// TIA Portal project "e045002v087-088" (V13) (continued)
VERSION : 0.1
// stored: InstanceOfName FB_CTR_VAL
"FB_CTR_VAL"
BEGIN
END_DATA_BLOCK

DATA_BLOCK "STOP_PALLET"   // DB78
{ S7_Optimized_Access := 'FALSE' }
VERSION : 0.1
// stored: InstanceOfName FB_CTR_VAL
"FB_CTR_VAL"
BEGIN
END_DATA_BLOCK

DATA_BLOCK "FB_CTR_MOT_FRD_DB"   // DB104
{ S7_Optimized_Access := 'FALSE' }
VERSION : 0.1
// stored: InstanceOfName FB_CTR_MOT_FRD
"FB_CTR_MOT_FRD"
BEGIN
END_DATA_BLOCK

DATA_BLOCK "FB_CTR_MOT_FRD_DB_1"   // DB109
{ S7_Optimized_Access := 'FALSE' }
VERSION : 0.1
// stored: InstanceOfName FB_CTR_MOT_FRD
"FB_CTR_MOT_FRD"
BEGIN
END_DATA_BLOCK

DATA_BLOCK "FB_CTR_MOT_FRD_DB_2"   // DB145
{ S7_Optimized_Access := 'FALSE' }
VERSION : 0.1
// stored: InstanceOfName FB_CTR_MOT_FRD
"FB_CTR_MOT_FRD"
BEGIN
END_DATA_BLOCK

// folder: Movimiento DATOS

DATA_BLOCK "DB_RECETAS"   // DB4
{ S7_Optimized_Access := 'FALSE' }
VERSION : 0.1
   VAR
      Receta : Array [1..10] of "Recetas";
      Static_1 : Bool;
   END_VAR
BEGIN
END_DATA_BLOCK

DATA_BLOCK "Puntero"   // DB7
{ S7_Optimized_Access := 'FALSE' }
VERSION : 0.1
   VAR
      Max_Nro_Elementos : Word;
      Max_Nro_Filas : Word;
      Max_Nro_Capas : Word;
      Max_Nro_Recetas : Word;
      Offset_Filas_HMI : Word;
      Length_Filas_HMI : Word;
      Offset_Elementos_HMI : Word;
      Length_Elementos_HMI : Word;
      Offset_Recetas : Word;
      Length_Recetas : Word;
      Offset_Nombre_Receta : Word;
      Length_Nombre_Receta : Word;
      Offset_CantCapas_Receta : Word;
      Offset_CapasDist_Receta : Word;
      Offset_Capas_Receta : Word;
      Length_Capas_Receta : Word;
      Offset_Filas_CapaReceta : Word;
      Length_Filas_CapaReceta : Word;
      Offset_Vel_Dosificador : Word;
      Length_Vel_Dosificador : Word;
   END_VAR
BEGIN
END_DATA_BLOCK

DATA_BLOCK "DB_Receta_Actual"   // DB42
{ S7_Optimized_Access := 'FALSE' }
VERSION : 0.1
   VAR
      Número : Byte;
      Nombre : Array [1 .. 50] of Char;
      Nro_Capas_Pallet : Byte;
      Nro_Capas_Distintas : Byte;
      Capa : Array [1..10] of "Capas_Proceso";
      Static_1 : Bool;
   END_VAR
BEGIN
END_DATA_BLOCK

// folder: (top level)

FUNCTION "Valida_Velocidades" : Void   // FC2, LAD
{ S7_Optimized_Access := 'FALSE' }
VERSION : 0.1
BEGIN

REGION Network 1: Dosificador
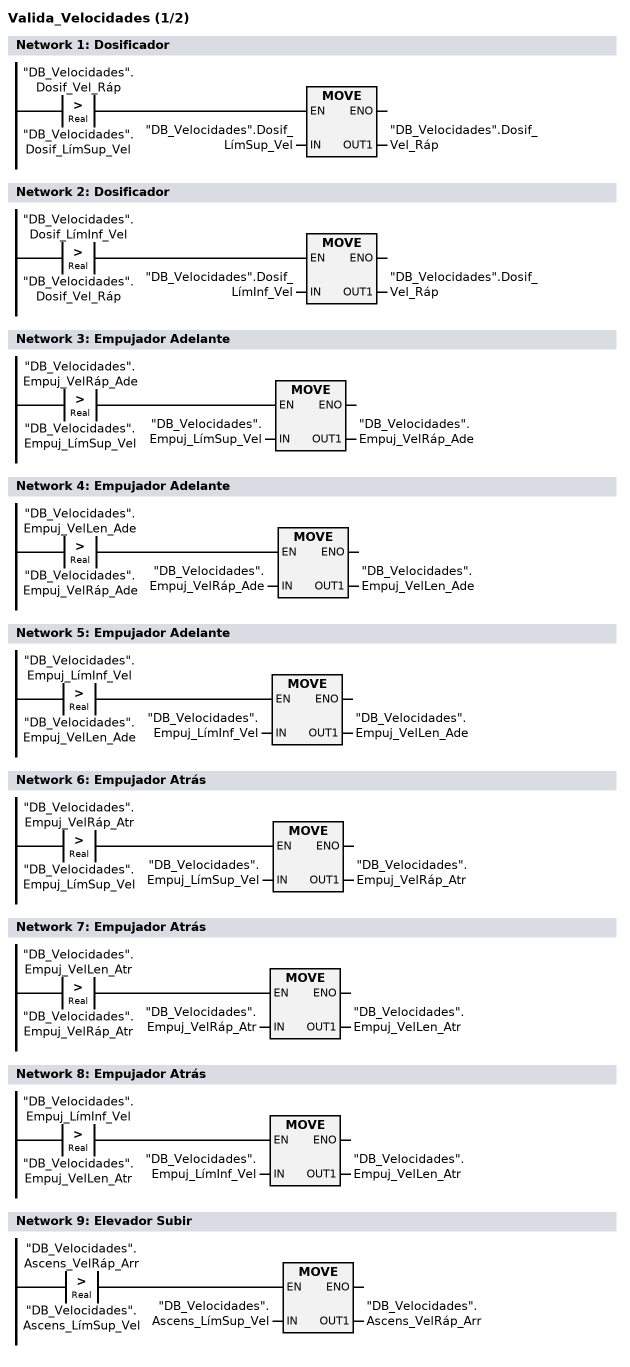
   RUNG wire#powerrail
      { S7_Templates := "SrcType := Real" } GT_Contact(in1 := "DB_Velocidades".Dosif_Vel_Ráp, in2 := "DB_Velocidades".Dosif_LímSup_Vel)
      { S7_GenerateENO := "TRUE" } Move(in := "DB_Velocidades".Dosif_LímSup_Vel, out1 => "DB_Velocidades".Dosif_Vel_Ráp)
   END_RUNG
   // the same network as SCL:
   IF "DB_Velocidades".Dosif_Vel_Ráp > "DB_Velocidades".Dosif_LímSup_Vel THEN
       "DB_Velocidades".Dosif_Vel_Ráp := "DB_Velocidades".Dosif_LímSup_Vel;
   END_IF;
END_REGION

REGION Network 2: Dosificador
   RUNG wire#powerrail
      { S7_Templates := "SrcType := Real" } GT_Contact(in1 := "DB_Velocidades".Dosif_LímInf_Vel, in2 := "DB_Velocidades".Dosif_Vel_Ráp)
      { S7_GenerateENO := "TRUE" } Move(in := "DB_Velocidades".Dosif_LímInf_Vel, out1 => "DB_Velocidades".Dosif_Vel_Ráp)
   END_RUNG
   // the same network as SCL:
   IF "DB_Velocidades".Dosif_LímInf_Vel > "DB_Velocidades".Dosif_Vel_Ráp THEN
       "DB_Velocidades".Dosif_Vel_Ráp := "DB_Velocidades".Dosif_LímInf_Vel;
   END_IF;
END_REGION

REGION Network 3: Empujador Adelante
   RUNG wire#powerrail
      { S7_Templates := "SrcType := Real" } GT_Contact(in1 := "DB_Velocidades".Empuj_VelRáp_Ade, in2 := "DB_Velocidades".Empuj_LímSup_Vel)
      { S7_GenerateENO := "TRUE" } Move(in := "DB_Velocidades".Empuj_LímSup_Vel, out1 => "DB_Velocidades".Empuj_VelRáp_Ade)
   END_RUNG
   // the same network as SCL:
   IF "DB_Velocidades".Empuj_VelRáp_Ade > "DB_Velocidades".Empuj_LímSup_Vel THEN
       "DB_Velocidades".Empuj_VelRáp_Ade := "DB_Velocidades".Empuj_LímSup_Vel;
   END_IF;
END_REGION

REGION Network 4: Empujador Adelante
   RUNG wire#powerrail
      { S7_Templates := "SrcType := Real" } GT_Contact(in1 := "DB_Velocidades".Empuj_VelLen_Ade, in2 := "DB_Velocidades".Empuj_VelRáp_Ade)
      { S7_GenerateENO := "TRUE" } Move(in := "DB_Velocidades".Empuj_VelRáp_Ade, out1 => "DB_Velocidades".Empuj_VelLen_Ade)
   END_RUNG
   // the same network as SCL:
   IF "DB_Velocidades".Empuj_VelLen_Ade > "DB_Velocidades".Empuj_VelRáp_Ade THEN
       "DB_Velocidades".Empuj_VelLen_Ade := "DB_Velocidades".Empuj_VelRáp_Ade;
   END_IF;
END_REGION

REGION Network 5: Empujador Adelante
   RUNG wire#powerrail
      { S7_Templates := "SrcType := Real" } GT_Contact(in1 := "DB_Velocidades".Empuj_LímInf_Vel, in2 := "DB_Velocidades".Empuj_VelLen_Ade)
      { S7_GenerateENO := "TRUE" } Move(in := "DB_Velocidades".Empuj_LímInf_Vel, out1 => "DB_Velocidades".Empuj_VelLen_Ade)
   END_RUNG
   // the same network as SCL:
   IF "DB_Velocidades".Empuj_LímInf_Vel > "DB_Velocidades".Empuj_VelLen_Ade THEN
       "DB_Velocidades".Empuj_VelLen_Ade := "DB_Velocidades".Empuj_LímInf_Vel;
   END_IF;
END_REGION

REGION Network 6: Empujador Atrás
   RUNG wire#powerrail
      { S7_Templates := "SrcType := Real" } GT_Contact(in1 := "DB_Velocidades".Empuj_VelRáp_Atr, in2 := "DB_Velocidades".Empuj_LímSup_Vel)
      { S7_GenerateENO := "TRUE" } Move(in := "DB_Velocidades".Empuj_LímSup_Vel, out1 => "DB_Velocidades".Empuj_VelRáp_Atr)
   END_RUNG
   // the same network as SCL:
   IF "DB_Velocidades".Empuj_VelRáp_Atr > "DB_Velocidades".Empuj_LímSup_Vel THEN
       "DB_Velocidades".Empuj_VelRáp_Atr := "DB_Velocidades".Empuj_LímSup_Vel;
   END_IF;
END_REGION

REGION Network 7: Empujador Atrás
   RUNG wire#powerrail
      { S7_Templates := "SrcType := Real" } GT_Contact(in1 := "DB_Velocidades".Empuj_VelLen_Atr, in2 := "DB_Velocidades".Empuj_VelRáp_Atr)
      { S7_GenerateENO := "TRUE" } Move(in := "DB_Velocidades".Empuj_VelRáp_Atr, out1 => "DB_Velocidades".Empuj_VelLen_Atr)
   END_RUNG
   // the same network as SCL:
   IF "DB_Velocidades".Empuj_VelLen_Atr > "DB_Velocidades".Empuj_VelRáp_Atr THEN
       "DB_Velocidades".Empuj_VelLen_Atr := "DB_Velocidades".Empuj_VelRáp_Atr;
   END_IF;
END_REGION

REGION Network 8: Empujador Atrás
   RUNG wire#powerrail
      { S7_Templates := "SrcType := Real" } GT_Contact(in1 := "DB_Velocidades".Empuj_LímInf_Vel, in2 := "DB_Velocidades".Empuj_VelLen_Atr)
      { S7_GenerateENO := "TRUE" } Move(in := "DB_Velocidades".Empuj_LímInf_Vel, out1 => "DB_Velocidades".Empuj_VelLen_Atr)
   END_RUNG
   // the same network as SCL:
   IF "DB_Velocidades".Empuj_LímInf_Vel > "DB_Velocidades".Empuj_VelLen_Atr THEN
       "DB_Velocidades".Empuj_VelLen_Atr := "DB_Velocidades".Empuj_LímInf_Vel;
   END_IF;
END_REGION

REGION Network 9: Elevador Subir
   RUNG wire#powerrail
      { S7_Templates := "SrcType := Real" } GT_Contact(in1 := "DB_Velocidades".Ascens_VelRáp_Arr, in2 := "DB_Velocidades".Ascens_LímSup_Vel)
      { S7_GenerateENO := "TRUE" } Move(in := "DB_Velocidades".Ascens_LímSup_Vel, out1 => "DB_Velocidades".Ascens_VelRáp_Arr)
   END_RUNG
   // the same network as SCL:
   IF "DB_Velocidades".Ascens_VelRáp_Arr > "DB_Velocidades".Ascens_LímSup_Vel THEN
       "DB_Velocidades".Ascens_VelRáp_Arr := "DB_Velocidades".Ascens_LímSup_Vel;
   END_IF;
END_REGION

REGION Network 10: Elevador Subir
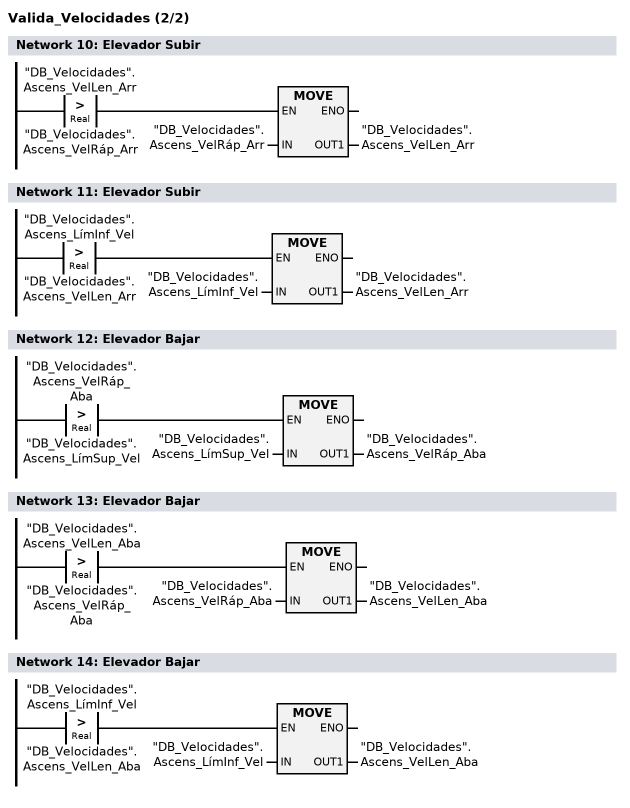
   RUNG wire#powerrail
      { S7_Templates := "SrcType := Real" } GT_Contact(in1 := "DB_Velocidades".Ascens_VelLen_Arr, in2 := "DB_Velocidades".Ascens_VelRáp_Arr)
      { S7_GenerateENO := "TRUE" } Move(in := "DB_Velocidades".Ascens_VelRáp_Arr, out1 => "DB_Velocidades".Ascens_VelLen_Arr)
   END_RUNG
   // the same network as SCL:
   IF "DB_Velocidades".Ascens_VelLen_Arr > "DB_Velocidades".Ascens_VelRáp_Arr THEN
       "DB_Velocidades".Ascens_VelLen_Arr := "DB_Velocidades".Ascens_VelRáp_Arr;
   END_IF;
END_REGION

REGION Network 11: Elevador Subir
   RUNG wire#powerrail
      { S7_Templates := "SrcType := Real" } GT_Contact(in1 := "DB_Velocidades".Ascens_LímInf_Vel, in2 := "DB_Velocidades".Ascens_VelLen_Arr)
      { S7_GenerateENO := "TRUE" } Move(in := "DB_Velocidades".Ascens_LímInf_Vel, out1 => "DB_Velocidades".Ascens_VelLen_Arr)
   END_RUNG
   // the same network as SCL:
   IF "DB_Velocidades".Ascens_LímInf_Vel > "DB_Velocidades".Ascens_VelLen_Arr THEN
       "DB_Velocidades".Ascens_VelLen_Arr := "DB_Velocidades".Ascens_LímInf_Vel;
   END_IF;
END_REGION

REGION Network 12: Elevador Bajar
   RUNG wire#powerrail
      { S7_Templates := "SrcType := Real" } GT_Contact(in1 := "DB_Velocidades".Ascens_VelRáp_Aba, in2 := "DB_Velocidades".Ascens_LímSup_Vel)
      { S7_GenerateENO := "TRUE" } Move(in := "DB_Velocidades".Ascens_LímSup_Vel, out1 => "DB_Velocidades".Ascens_VelRáp_Aba)
   END_RUNG
   // the same network as SCL:
   IF "DB_Velocidades".Ascens_VelRáp_Aba > "DB_Velocidades".Ascens_LímSup_Vel THEN
       "DB_Velocidades".Ascens_VelRáp_Aba := "DB_Velocidades".Ascens_LímSup_Vel;
   END_IF;
END_REGION

REGION Network 13: Elevador Bajar
   RUNG wire#powerrail
      { S7_Templates := "SrcType := Real" } GT_Contact(in1 := "DB_Velocidades".Ascens_VelLen_Aba, in2 := "DB_Velocidades".Ascens_VelRáp_Aba)
      { S7_GenerateENO := "TRUE" } Move(in := "DB_Velocidades".Ascens_VelRáp_Aba, out1 => "DB_Velocidades".Ascens_VelLen_Aba)
   END_RUNG
   // the same network as SCL:
   IF "DB_Velocidades".Ascens_VelLen_Aba > "DB_Velocidades".Ascens_VelRáp_Aba THEN
       "DB_Velocidades".Ascens_VelLen_Aba := "DB_Velocidades".Ascens_VelRáp_Aba;
   END_IF;
END_REGION

REGION Network 14: Elevador Bajar
   RUNG wire#powerrail
      { S7_Templates := "SrcType := Real" } GT_Contact(in1 := "DB_Velocidades".Ascens_LímInf_Vel, in2 := "DB_Velocidades".Ascens_VelLen_Aba)
      { S7_GenerateENO := "TRUE" } Move(in := "DB_Velocidades".Ascens_LímInf_Vel, out1 => "DB_Velocidades".Ascens_VelLen_Aba)
   END_RUNG
   // the same network as SCL:
   IF "DB_Velocidades".Ascens_LímInf_Vel > "DB_Velocidades".Ascens_VelLen_Aba THEN
       "DB_Velocidades".Ascens_VelLen_Aba := "DB_Velocidades".Ascens_LímInf_Vel;
   END_IF;
END_REGION
END_FUNCTION

FUNCTION "Genera_Flancos" : Void   // FC4, LAD
TITLE = Activa todos los flancos del programa
{ S7_Optimized_Access := 'FALSE' }
VERSION : 0.1
   VAR_TEMP   // added for the SCL form of the ladder/FBD networks
      _w1 : Bool;
      _w2 : Bool;
   END_VAR
BEGIN

REGION Network 1: "f"."nHMI.Pls_Inc_Elem"
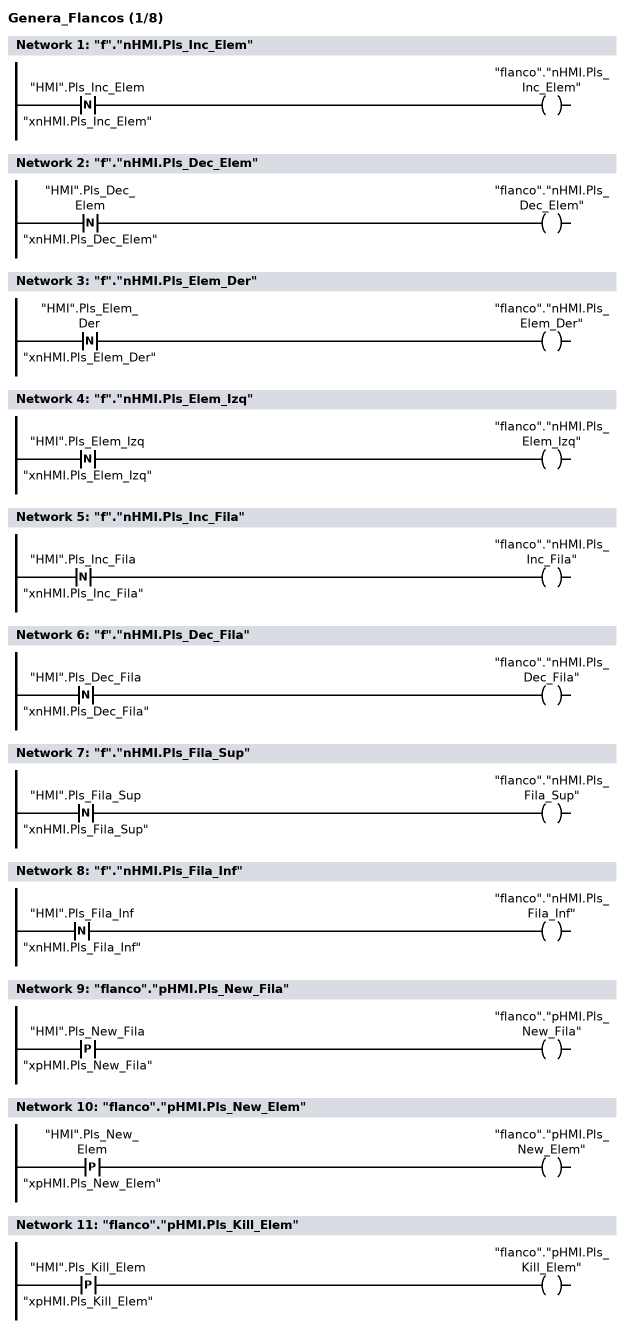
   RUNG wire#powerrail
      N_Contact(operand := "HMI".Pls_Inc_Elem, bit := "xnHMI.Pls_Inc_Elem")
      Coil( "flanco"."nHMI.Pls_Inc_Elem" )
   END_RUNG
   // the same network as SCL:
   #_w1 := NOT "HMI".Pls_Inc_Elem AND "xnHMI.Pls_Inc_Elem";   // falling edge of "HMI".Pls_Inc_Elem
   "xnHMI.Pls_Inc_Elem" := "HMI".Pls_Inc_Elem;
   "flanco"."nHMI.Pls_Inc_Elem" := #_w1;
END_REGION

REGION Network 2: "f"."nHMI.Pls_Dec_Elem"
   RUNG wire#powerrail
      N_Contact(operand := "HMI".Pls_Dec_Elem, bit := "xnHMI.Pls_Dec_Elem")
      Coil( "flanco"."nHMI.Pls_Dec_Elem" )
   END_RUNG
   // the same network as SCL:
   #_w1 := NOT "HMI".Pls_Dec_Elem AND "xnHMI.Pls_Dec_Elem";   // falling edge of "HMI".Pls_Dec_Elem
   "xnHMI.Pls_Dec_Elem" := "HMI".Pls_Dec_Elem;
   "flanco"."nHMI.Pls_Dec_Elem" := #_w1;
END_REGION

REGION Network 3: "f"."nHMI.Pls_Elem_Der"
   RUNG wire#powerrail
      N_Contact(operand := "HMI".Pls_Elem_Der, bit := "xnHMI.Pls_Elem_Der")
      Coil( "flanco"."nHMI.Pls_Elem_Der" )
   END_RUNG
   // the same network as SCL:
   #_w1 := NOT "HMI".Pls_Elem_Der AND "xnHMI.Pls_Elem_Der";   // falling edge of "HMI".Pls_Elem_Der
   "xnHMI.Pls_Elem_Der" := "HMI".Pls_Elem_Der;
   "flanco"."nHMI.Pls_Elem_Der" := #_w1;
END_REGION

REGION Network 4: "f"."nHMI.Pls_Elem_Izq"
   RUNG wire#powerrail
      N_Contact(operand := "HMI".Pls_Elem_Izq, bit := "xnHMI.Pls_Elem_Izq")
      Coil( "flanco"."nHMI.Pls_Elem_Izq" )
   END_RUNG
   // the same network as SCL:
   #_w1 := NOT "HMI".Pls_Elem_Izq AND "xnHMI.Pls_Elem_Izq";   // falling edge of "HMI".Pls_Elem_Izq
   "xnHMI.Pls_Elem_Izq" := "HMI".Pls_Elem_Izq;
   "flanco"."nHMI.Pls_Elem_Izq" := #_w1;
END_REGION

REGION Network 5: "f"."nHMI.Pls_Inc_Fila"
   RUNG wire#powerrail
      N_Contact(operand := "HMI".Pls_Inc_Fila, bit := "xnHMI.Pls_Inc_Fila")
      Coil( "flanco"."nHMI.Pls_Inc_Fila" )
   END_RUNG
   // the same network as SCL:
   #_w1 := NOT "HMI".Pls_Inc_Fila AND "xnHMI.Pls_Inc_Fila";   // falling edge of "HMI".Pls_Inc_Fila
   "xnHMI.Pls_Inc_Fila" := "HMI".Pls_Inc_Fila;
   "flanco"."nHMI.Pls_Inc_Fila" := #_w1;
END_REGION

REGION Network 6: "f"."nHMI.Pls_Dec_Fila"
   RUNG wire#powerrail
      N_Contact(operand := "HMI".Pls_Dec_Fila, bit := "xnHMI.Pls_Dec_Fila")
      Coil( "flanco"."nHMI.Pls_Dec_Fila" )
   END_RUNG
   // the same network as SCL:
   #_w1 := NOT "HMI".Pls_Dec_Fila AND "xnHMI.Pls_Dec_Fila";   // falling edge of "HMI".Pls_Dec_Fila
   "xnHMI.Pls_Dec_Fila" := "HMI".Pls_Dec_Fila;
   "flanco"."nHMI.Pls_Dec_Fila" := #_w1;
END_REGION

REGION Network 7: "f"."nHMI.Pls_Fila_Sup"
   RUNG wire#powerrail
      N_Contact(operand := "HMI".Pls_Fila_Sup, bit := "xnHMI.Pls_Fila_Sup")
      Coil( "flanco"."nHMI.Pls_Fila_Sup" )
   END_RUNG
   // the same network as SCL:
   #_w1 := NOT "HMI".Pls_Fila_Sup AND "xnHMI.Pls_Fila_Sup";   // falling edge of "HMI".Pls_Fila_Sup
   "xnHMI.Pls_Fila_Sup" := "HMI".Pls_Fila_Sup;
   "flanco"."nHMI.Pls_Fila_Sup" := #_w1;
END_REGION

REGION Network 8: "f"."nHMI.Pls_Fila_Inf"
   RUNG wire#powerrail
      N_Contact(operand := "HMI".Pls_Fila_Inf, bit := "xnHMI.Pls_Fila_Inf")
      Coil( "flanco"."nHMI.Pls_Fila_Inf" )
   END_RUNG
   // the same network as SCL:
   #_w1 := NOT "HMI".Pls_Fila_Inf AND "xnHMI.Pls_Fila_Inf";   // falling edge of "HMI".Pls_Fila_Inf
   "xnHMI.Pls_Fila_Inf" := "HMI".Pls_Fila_Inf;
   "flanco"."nHMI.Pls_Fila_Inf" := #_w1;
END_REGION

REGION Network 9: "flanco"."pHMI.Pls_New_Fila"
   RUNG wire#powerrail
      P_Contact(operand := "HMI".Pls_New_Fila, bit := "xpHMI.Pls_New_Fila")
      Coil( "flanco"."pHMI.Pls_New_Fila" )
   END_RUNG
   // the same network as SCL:
   #_w1 := "HMI".Pls_New_Fila AND NOT "xpHMI.Pls_New_Fila";   // rising edge of "HMI".Pls_New_Fila
   "xpHMI.Pls_New_Fila" := "HMI".Pls_New_Fila;
   "flanco"."pHMI.Pls_New_Fila" := #_w1;
END_REGION

REGION Network 10: "flanco"."pHMI.Pls_New_Elem"
   RUNG wire#powerrail
      P_Contact(operand := "HMI".Pls_New_Elem, bit := "xpHMI.Pls_New_Elem")
      Coil( "flanco"."pHMI.Pls_New_Elem" )
   END_RUNG
   // the same network as SCL:
   #_w1 := "HMI".Pls_New_Elem AND NOT "xpHMI.Pls_New_Elem";   // rising edge of "HMI".Pls_New_Elem
   "xpHMI.Pls_New_Elem" := "HMI".Pls_New_Elem;
   "flanco"."pHMI.Pls_New_Elem" := #_w1;
END_REGION

REGION Network 11: "flanco"."pHMI.Pls_Kill_Elem"
   RUNG wire#powerrail
      P_Contact(operand := "HMI".Pls_Kill_Elem, bit := "xpHMI.Pls_Kill_Elem")
      Coil( "flanco"."pHMI.Pls_Kill_Elem" )
   END_RUNG
   // the same network as SCL:
   #_w1 := "HMI".Pls_Kill_Elem AND NOT "xpHMI.Pls_Kill_Elem";   // rising edge of "HMI".Pls_Kill_Elem
   "xpHMI.Pls_Kill_Elem" := "HMI".Pls_Kill_Elem;
   "flanco"."pHMI.Pls_Kill_Elem" := #_w1;
END_REGION

REGION Network 12: "f"."nHMI.Pls_WR_Receta"
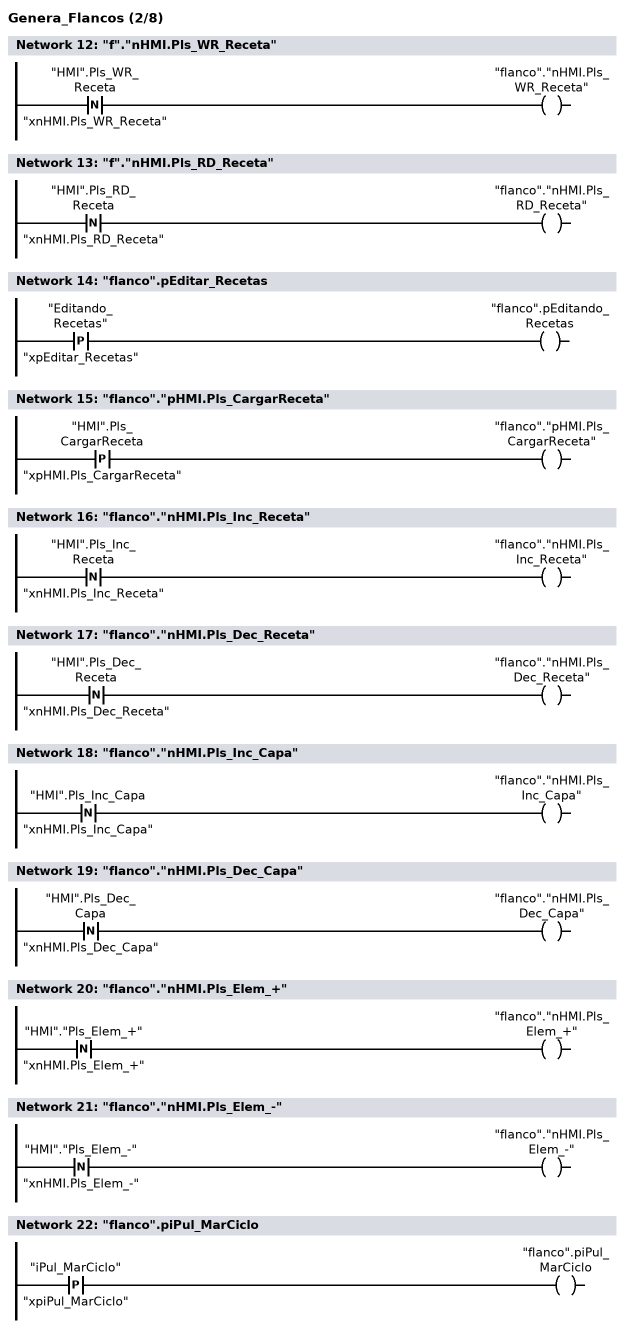
   RUNG wire#powerrail
      N_Contact(operand := "HMI".Pls_WR_Receta, bit := "xnHMI.Pls_WR_Receta")
      Coil( "flanco"."nHMI.Pls_WR_Receta" )
   END_RUNG
   // the same network as SCL:
   #_w1 := NOT "HMI".Pls_WR_Receta AND "xnHMI.Pls_WR_Receta";   // falling edge of "HMI".Pls_WR_Receta
   "xnHMI.Pls_WR_Receta" := "HMI".Pls_WR_Receta;
   "flanco"."nHMI.Pls_WR_Receta" := #_w1;
END_REGION

REGION Network 13: "f"."nHMI.Pls_RD_Receta"
   RUNG wire#powerrail
      N_Contact(operand := "HMI".Pls_RD_Receta, bit := "xnHMI.Pls_RD_Receta")
      Coil( "flanco"."nHMI.Pls_RD_Receta" )
   END_RUNG
   // the same network as SCL:
   #_w1 := NOT "HMI".Pls_RD_Receta AND "xnHMI.Pls_RD_Receta";   // falling edge of "HMI".Pls_RD_Receta
   "xnHMI.Pls_RD_Receta" := "HMI".Pls_RD_Receta;
   "flanco"."nHMI.Pls_RD_Receta" := #_w1;
END_REGION

REGION Network 14: "flanco".pEditar_Recetas
   RUNG wire#powerrail
      P_Contact(operand := "Editando_Recetas", bit := "xpEditar_Recetas")
      Coil( "flanco".pEditando_Recetas )
   END_RUNG
   // the same network as SCL:
   #_w1 := "Editando_Recetas" AND NOT "xpEditar_Recetas";   // rising edge of "Editando_Recetas"
   "xpEditar_Recetas" := "Editando_Recetas";
   "flanco".pEditando_Recetas := #_w1;
END_REGION

REGION Network 15: "flanco"."pHMI.Pls_CargarReceta"
   RUNG wire#powerrail
      P_Contact(operand := "HMI".Pls_CargarReceta, bit := "xpHMI.Pls_CargarReceta")
      Coil( "flanco"."pHMI.Pls_CargarReceta" )
   END_RUNG
   // the same network as SCL:
   #_w1 := "HMI".Pls_CargarReceta AND NOT "xpHMI.Pls_CargarReceta";   // rising edge of "HMI".Pls_CargarReceta
   "xpHMI.Pls_CargarReceta" := "HMI".Pls_CargarReceta;
   "flanco"."pHMI.Pls_CargarReceta" := #_w1;
END_REGION

REGION Network 16: "flanco"."nHMI.Pls_Inc_Receta"
   RUNG wire#powerrail
      N_Contact(operand := "HMI".Pls_Inc_Receta, bit := "xnHMI.Pls_Inc_Receta")
      Coil( "flanco"."nHMI.Pls_Inc_Receta" )
   END_RUNG
   // the same network as SCL:
   #_w1 := NOT "HMI".Pls_Inc_Receta AND "xnHMI.Pls_Inc_Receta";   // falling edge of "HMI".Pls_Inc_Receta
   "xnHMI.Pls_Inc_Receta" := "HMI".Pls_Inc_Receta;
   "flanco"."nHMI.Pls_Inc_Receta" := #_w1;
END_REGION

REGION Network 17: "flanco"."nHMI.Pls_Dec_Receta"
   RUNG wire#powerrail
      N_Contact(operand := "HMI".Pls_Dec_Receta, bit := "xnHMI.Pls_Dec_Receta")
      Coil( "flanco"."nHMI.Pls_Dec_Receta" )
   END_RUNG
   // the same network as SCL:
   #_w1 := NOT "HMI".Pls_Dec_Receta AND "xnHMI.Pls_Dec_Receta";   // falling edge of "HMI".Pls_Dec_Receta
   "xnHMI.Pls_Dec_Receta" := "HMI".Pls_Dec_Receta;
   "flanco"."nHMI.Pls_Dec_Receta" := #_w1;
END_REGION

REGION Network 18: "flanco"."nHMI.Pls_Inc_Capa"
   RUNG wire#powerrail
      N_Contact(operand := "HMI".Pls_Inc_Capa, bit := "xnHMI.Pls_Inc_Capa")
      Coil( "flanco"."nHMI.Pls_Inc_Capa" )
   END_RUNG
   // the same network as SCL:
   #_w1 := NOT "HMI".Pls_Inc_Capa AND "xnHMI.Pls_Inc_Capa";   // falling edge of "HMI".Pls_Inc_Capa
   "xnHMI.Pls_Inc_Capa" := "HMI".Pls_Inc_Capa;
   "flanco"."nHMI.Pls_Inc_Capa" := #_w1;
END_REGION

REGION Network 19: "flanco"."nHMI.Pls_Dec_Capa"
   RUNG wire#powerrail
      N_Contact(operand := "HMI".Pls_Dec_Capa, bit := "xnHMI.Pls_Dec_Capa")
      Coil( "flanco"."nHMI.Pls_Dec_Capa" )
   END_RUNG
   // the same network as SCL:
   #_w1 := NOT "HMI".Pls_Dec_Capa AND "xnHMI.Pls_Dec_Capa";   // falling edge of "HMI".Pls_Dec_Capa
   "xnHMI.Pls_Dec_Capa" := "HMI".Pls_Dec_Capa;
   "flanco"."nHMI.Pls_Dec_Capa" := #_w1;
END_REGION

REGION Network 20: "flanco"."nHMI.Pls_Elem_+"
   RUNG wire#powerrail
      N_Contact(operand := "HMI"."Pls_Elem_+", bit := "xnHMI.Pls_Elem_+")
      Coil( "flanco"."nHMI.Pls_Elem_+" )
   END_RUNG
   // the same network as SCL:
   #_w1 := NOT "HMI"."Pls_Elem_+" AND "xnHMI.Pls_Elem_+";   // falling edge of "HMI"."Pls_Elem_+"
   "xnHMI.Pls_Elem_+" := "HMI"."Pls_Elem_+";
   "flanco"."nHMI.Pls_Elem_+" := #_w1;
END_REGION

REGION Network 21: "flanco"."nHMI.Pls_Elem_-"
   RUNG wire#powerrail
      N_Contact(operand := "HMI"."Pls_Elem_-", bit := "xnHMI.Pls_Elem_-")
      Coil( "flanco"."nHMI.Pls_Elem_-" )
   END_RUNG
   // the same network as SCL:
   #_w1 := NOT "HMI"."Pls_Elem_-" AND "xnHMI.Pls_Elem_-";   // falling edge of "HMI"."Pls_Elem_-"
   "xnHMI.Pls_Elem_-" := "HMI"."Pls_Elem_-";
   "flanco"."nHMI.Pls_Elem_-" := #_w1;
END_REGION

REGION Network 22: "flanco".piPul_MarCiclo
   RUNG wire#powerrail
      P_Contact(operand := "iPul_MarCiclo", bit := "xpiPul_MarCiclo")
      Coil( "flanco".piPul_MarCiclo )
   END_RUNG
   // the same network as SCL:
   #_w1 := "iPul_MarCiclo" AND NOT "xpiPul_MarCiclo";   // rising edge of "iPul_MarCiclo"
   "xpiPul_MarCiclo" := "iPul_MarCiclo";
   "flanco".piPul_MarCiclo := #_w1;
END_REGION

REGION Network 23: "flanco".piPul_HabTransp
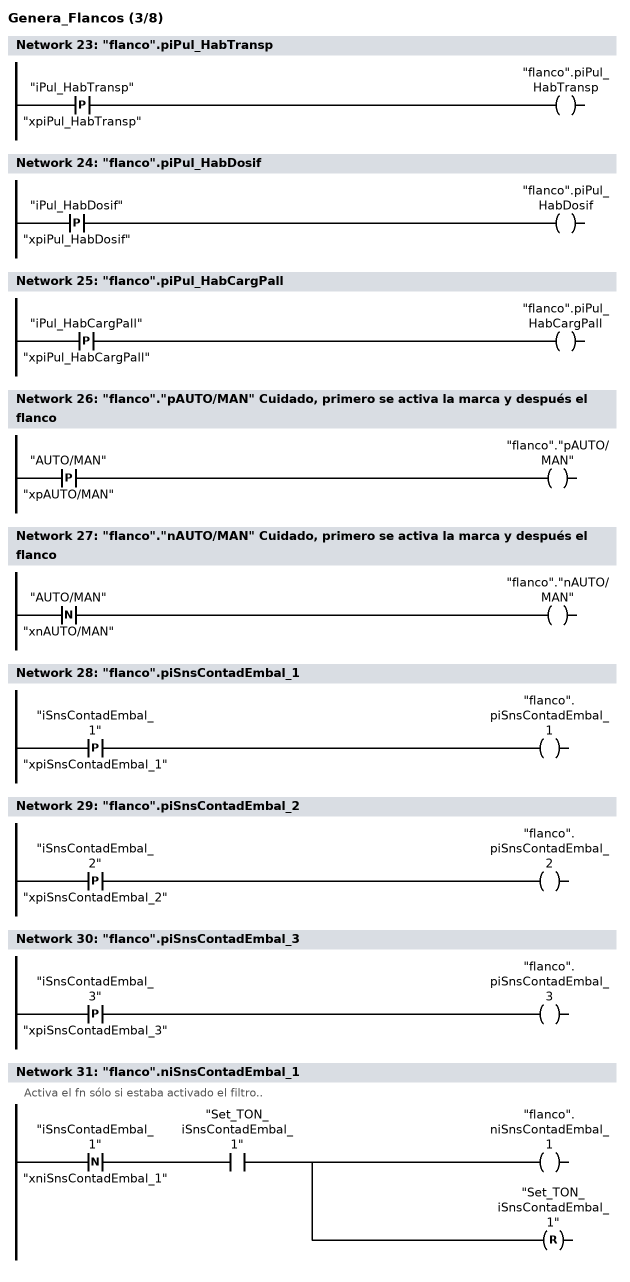
   RUNG wire#powerrail
      P_Contact(operand := "iPul_HabTransp", bit := "xpiPul_HabTransp")
      Coil( "flanco".piPul_HabTransp )
   END_RUNG
   // the same network as SCL:
   #_w1 := "iPul_HabTransp" AND NOT "xpiPul_HabTransp";   // rising edge of "iPul_HabTransp"
   "xpiPul_HabTransp" := "iPul_HabTransp";
   "flanco".piPul_HabTransp := #_w1;
END_REGION

REGION Network 24: "flanco".piPul_HabDosif
   RUNG wire#powerrail
      P_Contact(operand := "iPul_HabDosif", bit := "xpiPul_HabDosif")
      Coil( "flanco".piPul_HabDosif )
   END_RUNG
   // the same network as SCL:
   #_w1 := "iPul_HabDosif" AND NOT "xpiPul_HabDosif";   // rising edge of "iPul_HabDosif"
   "xpiPul_HabDosif" := "iPul_HabDosif";
   "flanco".piPul_HabDosif := #_w1;
END_REGION

REGION Network 25: "flanco".piPul_HabCargPall
   RUNG wire#powerrail
      P_Contact(operand := "iPul_HabCargPall", bit := "xpiPul_HabCargPall")
      Coil( "flanco".piPul_HabCargPall )
   END_RUNG
   // the same network as SCL:
   #_w1 := "iPul_HabCargPall" AND NOT "xpiPul_HabCargPall";   // rising edge of "iPul_HabCargPall"
   "xpiPul_HabCargPall" := "iPul_HabCargPall";
   "flanco".piPul_HabCargPall := #_w1;
END_REGION

REGION Network 26: "flanco"."pAUTO/MAN" Cuidado, primero se activa la marca y después el flanco
   RUNG wire#powerrail
      P_Contact(operand := "AUTO/MAN", bit := "xpAUTO/MAN")
      Coil( "flanco"."pAUTO/MAN" )
   END_RUNG
   // the same network as SCL:
   #_w1 := "AUTO/MAN" AND NOT "xpAUTO/MAN";   // rising edge of "AUTO/MAN"
   "xpAUTO/MAN" := "AUTO/MAN";
   "flanco"."pAUTO/MAN" := #_w1;
END_REGION

REGION Network 27: "flanco"."nAUTO/MAN" Cuidado, primero se activa la marca y después el flanco
   RUNG wire#powerrail
      N_Contact(operand := "AUTO/MAN", bit := "xnAUTO/MAN")
      Coil( "flanco"."nAUTO/MAN" )
   END_RUNG
   // the same network as SCL:
   #_w1 := NOT "AUTO/MAN" AND "xnAUTO/MAN";   // falling edge of "AUTO/MAN"
   "xnAUTO/MAN" := "AUTO/MAN";
   "flanco"."nAUTO/MAN" := #_w1;
END_REGION

REGION Network 28: "flanco".piSnsContadEmbal_1
   RUNG wire#powerrail
      P_Contact(operand := "iSnsContadEmbal_1", bit := "xpiSnsContadEmbal_1")
      Coil( "flanco".piSnsContadEmbal_1 )
   END_RUNG
   // the same network as SCL:
   #_w1 := "iSnsContadEmbal_1" AND NOT "xpiSnsContadEmbal_1";   // rising edge of "iSnsContadEmbal_1"
   "xpiSnsContadEmbal_1" := "iSnsContadEmbal_1";
   "flanco".piSnsContadEmbal_1 := #_w1;
END_REGION

REGION Network 29: "flanco".piSnsContadEmbal_2
   RUNG wire#powerrail
      P_Contact(operand := "iSnsContadEmbal_2", bit := "xpiSnsContadEmbal_2")
      Coil( "flanco".piSnsContadEmbal_2 )
   END_RUNG
   // the same network as SCL:
   #_w1 := "iSnsContadEmbal_2" AND NOT "xpiSnsContadEmbal_2";   // rising edge of "iSnsContadEmbal_2"
   "xpiSnsContadEmbal_2" := "iSnsContadEmbal_2";
   "flanco".piSnsContadEmbal_2 := #_w1;
END_REGION

REGION Network 30: "flanco".piSnsContadEmbal_3
   RUNG wire#powerrail
      P_Contact(operand := "iSnsContadEmbal_3", bit := "xpiSnsContadEmbal_3")
      Coil( "flanco".piSnsContadEmbal_3 )
   END_RUNG
   // the same network as SCL:
   #_w1 := "iSnsContadEmbal_3" AND NOT "xpiSnsContadEmbal_3";   // rising edge of "iSnsContadEmbal_3"
   "xpiSnsContadEmbal_3" := "iSnsContadEmbal_3";
   "flanco".piSnsContadEmbal_3 := #_w1;
END_REGION

REGION Network 31: "flanco".niSnsContadEmbal_1
   // Activa el fn sólo si estaba activado el filtro..
   RUNG wire#powerrail
      N_Contact(operand := "iSnsContadEmbal_1", bit := "xniSnsContadEmbal_1")
      Contact( "Set_TON_iSnsContadEmbal_1" )
      wire#w1
      Coil( "flanco".niSnsContadEmbal_1 )
   END_RUNG
   RUNG wire#w1
      R_Coil( "Set_TON_iSnsContadEmbal_1" )
   END_RUNG
   // the same network as SCL:
   #_w1 := NOT "iSnsContadEmbal_1" AND "xniSnsContadEmbal_1";   // falling edge of "iSnsContadEmbal_1"
   "xniSnsContadEmbal_1" := "iSnsContadEmbal_1";
   "flanco".niSnsContadEmbal_1 := #_w1 AND "Set_TON_iSnsContadEmbal_1";
   IF "flanco".niSnsContadEmbal_1 THEN "Set_TON_iSnsContadEmbal_1" := FALSE; END_IF;
END_REGION

REGION Network 32: "flanco".niSnsContadEmbal_2
   // Activa el fn sólo si estaba activado el filtro..
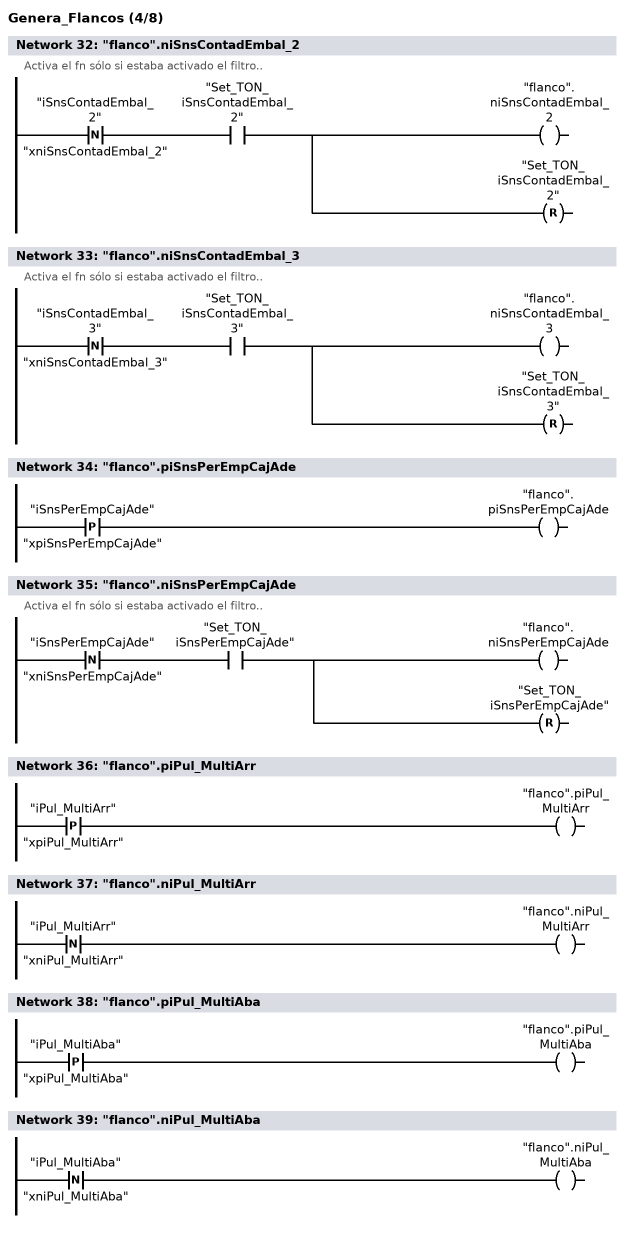
   RUNG wire#powerrail
      N_Contact(operand := "iSnsContadEmbal_2", bit := "xniSnsContadEmbal_2")
      Contact( "Set_TON_iSnsContadEmbal_2" )
      wire#w1
      Coil( "flanco".niSnsContadEmbal_2 )
   END_RUNG
   RUNG wire#w1
      R_Coil( "Set_TON_iSnsContadEmbal_2" )
   END_RUNG
   // the same network as SCL:
   #_w1 := NOT "iSnsContadEmbal_2" AND "xniSnsContadEmbal_2";   // falling edge of "iSnsContadEmbal_2"
   "xniSnsContadEmbal_2" := "iSnsContadEmbal_2";
   "flanco".niSnsContadEmbal_2 := #_w1 AND "Set_TON_iSnsContadEmbal_2";
   IF "flanco".niSnsContadEmbal_2 THEN "Set_TON_iSnsContadEmbal_2" := FALSE; END_IF;
END_REGION

REGION Network 33: "flanco".niSnsContadEmbal_3
   // Activa el fn sólo si estaba activado el filtro..
   RUNG wire#powerrail
      N_Contact(operand := "iSnsContadEmbal_3", bit := "xniSnsContadEmbal_3")
      Contact( "Set_TON_iSnsContadEmbal_3" )
      wire#w1
      Coil( "flanco".niSnsContadEmbal_3 )
   END_RUNG
   RUNG wire#w1
      R_Coil( "Set_TON_iSnsContadEmbal_3" )
   END_RUNG
   // the same network as SCL:
   #_w1 := NOT "iSnsContadEmbal_3" AND "xniSnsContadEmbal_3";   // falling edge of "iSnsContadEmbal_3"
   "xniSnsContadEmbal_3" := "iSnsContadEmbal_3";
   "flanco".niSnsContadEmbal_3 := #_w1 AND "Set_TON_iSnsContadEmbal_3";
   IF "flanco".niSnsContadEmbal_3 THEN "Set_TON_iSnsContadEmbal_3" := FALSE; END_IF;
END_REGION

REGION Network 34: "flanco".piSnsPerEmpCajAde
   RUNG wire#powerrail
      P_Contact(operand := "iSnsPerEmpCajAde", bit := "xpiSnsPerEmpCajAde")
      Coil( "flanco".piSnsPerEmpCajAde )
   END_RUNG
   // the same network as SCL:
   #_w1 := "iSnsPerEmpCajAde" AND NOT "xpiSnsPerEmpCajAde";   // rising edge of "iSnsPerEmpCajAde"
   "xpiSnsPerEmpCajAde" := "iSnsPerEmpCajAde";
   "flanco".piSnsPerEmpCajAde := #_w1;
END_REGION

REGION Network 35: "flanco".niSnsPerEmpCajAde
   // Activa el fn sólo si estaba activado el filtro..
   RUNG wire#powerrail
      N_Contact(operand := "iSnsPerEmpCajAde", bit := "xniSnsPerEmpCajAde")
      Contact( "Set_TON_iSnsPerEmpCajAde" )
      wire#w1
      Coil( "flanco".niSnsPerEmpCajAde )
   END_RUNG
   RUNG wire#w1
      R_Coil( "Set_TON_iSnsPerEmpCajAde" )
   END_RUNG
   // the same network as SCL:
   #_w1 := NOT "iSnsPerEmpCajAde" AND "xniSnsPerEmpCajAde";   // falling edge of "iSnsPerEmpCajAde"
   "xniSnsPerEmpCajAde" := "iSnsPerEmpCajAde";
   "flanco".niSnsPerEmpCajAde := #_w1 AND "Set_TON_iSnsPerEmpCajAde";
   IF "flanco".niSnsPerEmpCajAde THEN "Set_TON_iSnsPerEmpCajAde" := FALSE; END_IF;
END_REGION

REGION Network 36: "flanco".piPul_MultiArr
   RUNG wire#powerrail
      P_Contact(operand := "iPul_MultiArr", bit := "xpiPul_MultiArr")
      Coil( "flanco".piPul_MultiArr )
   END_RUNG
   // the same network as SCL:
   #_w1 := "iPul_MultiArr" AND NOT "xpiPul_MultiArr";   // rising edge of "iPul_MultiArr"
   "xpiPul_MultiArr" := "iPul_MultiArr";
   "flanco".piPul_MultiArr := #_w1;
END_REGION

